             //Try reconnection after a wait time
             #statIterator := 0;
             #statState.connection := #STATE_WAIT;
           END_IF;
         END_IF;
         //Job completed without error
       ELSIF (#instTCON.DONE) THEN

         //Connection successfully established
         #diagnostics.statistics.totalReconnects := #diagnostics.statistics.totalReconnects + 1;
         #statState.connection := #OPERATION;

         #error := FALSE;

         //Reset all state machines
         #statState.receiver := #READ;
         #statState.sender := #STATE_INACTIVE;
         #statState.comReceiver := #LCOM_EXPECTED;
         #statState.comSender := #STATE_INACTIVE;
         //Receive
         #statReceive.trcvFct.dataOffset := 0;
         #statReceive.trcvFct.dataLength := 0;
         #statReceive.trcvFct.dataLengthRest := 0;
         #statReceive.trcvFct.dataReceived := FALSE;
         #statReceive.tempTelegram.index := 0;
         #statReceive.tempTelegram.telegramType := 0;
         #statReceive.numberOfLComHeader := 0;
         #statReceive.dataTelegram.totalMessageLength := 0;
         #statReceive.dataTelegram.actPackageLength := 0;
         #statReceive.dataTelegram.ackMessageOffset := 0;
         #statReceive.dataTelegram.messageOffset := 0;
         #statReceive.dataTelegram.ackMessageCounter := 0;
         #statReceive.dataTelegram.messageCounter := 0;
         #statReceive.userData.totalLength := 0;
         #statReceive.userData.offset := 0;
         //Send
         #statSend.tsendFct.dataLengthRest := 0;
         #statSend.tsendFct.dataOffset := 0;
         #statSend.tsendFct.status := 16#0000;
         #statSend.expectedAck.package1.offset := 0;
         #statSend.dataTelegram.messageCounter := 0;
         #statSend.dataTelegram.ackMessageCounter := 0;
         #statSend.dataTelegram.messageOffset := 0;
         #statSend.dataTelegram.ackMessageOffset := 0;
         #statSend.dataTelegram.actPackageLength := 0;
         #statSend.dataTelegram.totalMessageLength := 0;
         #statSend.numberOfLComPackage := 0;
         #statSend.userData.totalLength := 0;
         #statSend.userData.offset := 0;
         #statSend.userData.sendCycleViolation := FALSE;
         #statOldSend := FALSE;

         #diagnostics.statistics.maxMsgSendingTime := T#0ms;
         #diagnostics.localConfig.sender.cycleTime := T#0ms;
         #diagnostics.localConfig.sender.ackTimeout := T#0ms;

         #diagnostics.statistics.lastTimeSync.YEAR := 2200;
         #statCopyNBytes := 0;

         //Reset all timer
         #instLocalLifeSignCycleTimer(IN := FALSE,
                                      PT := #diagnostics.localConfig.connection.lifeSignCycleTime);

         #instPartnerLifeSignCycleTimer(IN := FALSE,
                                        PT := (#diagnostics.partnerConfig.connnection.lifeSignCycleTime));

         #instLocalCycleTimeTimer(IN := FALSE,
                                  PT := #diagnostics.localConfig.sender.cycleTime);

         #instExpectedAckPackage1(IN := FALSE,
                                  PT := #diagnostics.localConfig.sender.ackTimeout);

         #instSyncTimer(IN := FALSE,
                        PT := T#1s);

         #instSendErrorTimer(IN := FALSE,
                             PT := #MAX_TRIAL_TIME);

         #instRcvErrorTimer(IN := FALSE,
                            PT := #MAX_TRIAL_TIME);

         //Reset all active failures in the diagnostics buffer
         FOR #statIterator := 0 TO #DIAG_BUFFER_UPPER_LIM BY 1 DO
           #diagnostics.buffer[#statIterator].isActive := FALSE;
         END_FOR;

         //With LCom protocol
         IF (#diagnostics.localConfig.connection.useLComProtocol = TRUE) THEN

           IF (#statConnectAttempts MOD 2 = 0) THEN
             //1st try LCom Version 2.0
             #statActualLocalLComVersion := #LCOM_HEADER_V2;
             #statSend.configTelegramV2.LComVersion := #LCOM_HEADER_V2;
             #statSend.configTelegramV2.status := BOOL_TO_BYTE(#diagnostics.localConfig.timeSync.usePartnerTimestamps);
             #statSend.configTelegramV2.sendModeSyncTime := #diagnostics.localConfig.timeSync.sendMode;
             #statSend.configTelegramV2.lifeSignCycle := #diagnostics.localConfig.connection.lifeSignCycleTime;
             #statSend.configTelegramV2.cycleTime := #configuration.sender.cycleTime;
             #statSend.configTelegramV2.ackTimeOut := #configuration.sender.ackTimeout;
             #statSend.configTelegramV2.maxSendDataLength := #diagnostics.localConfig.sizeOfSendBuffer;
             #statSend.configTelegramV2.maxReceiveDataLength := #diagnostics.localConfig.sizeOfReceiveBuffer;

             #statSend.dataTelegram.LComVersion := #statSend.configTelegramV2.LComVersion;
           ELSE
             //2nd try LCom Version 1.0
             #statActualLocalLComVersion := #LCOM_HEADER_V1;
             #statSend.configTelegramV1.LComVersion := #LCOM_HEADER_V1;
             #statSend.configTelegramV1.comMode := 16#03;
             #statSend.configTelegramV1.slidingWindow := 1;
             #statSend.configTelegramV1.status := BOOL_TO_BYTE(#diagnostics.localConfig.timeSync.usePartnerTimestamps);
             #statSend.configTelegramV1.sendModeSyncTime := #diagnostics.localConfig.timeSync.sendMode;

             #statSend.dataTelegram.LComVersion := #statSend.configTelegramV1.LComVersion;

             //Check max. lifeSignCycleTime
             IF (#diagnostics.localConfig.connection.lifeSignCycleTime > T#65535ms) THEN

               #statDiag.bufferIndex := #statDiag.bufferIndex + 1;
               #statDiag.buffer[#statDiag.bufferIndex].additionalValue4 := #diagnostics.localConfig.connection.lifeSignCycleTime;
               #diagnostics.localConfig.connection.lifeSignCycleTime := T#65535ms;

               #statDiag.buffer[#statDiag.bufferIndex].status := "LCOM_WARN_LIFE_SIGN_LIMITATION";
               #statDiag.buffer[#statDiag.bufferIndex].subFunctionErrorID := 16#0000;
               #statDiag.buffer[#statDiag.bufferIndex].additionalValue1 := 65535.0;
               #statDiag.buffer[#statDiag.bufferIndex].additionalValue2 := 0.0;
               #statDiag.buffer[#statDiag.bufferIndex].additionalValue3 := 0.0;
             ELSE
               ;
             END_IF;
             #statSend.configTelegramV1.lifeSignCycle := TIME_TO_UINT(#diagnostics.localConfig.connection.lifeSignCycleTime);

             //Check max.sizeOfSendBuffer
             IF (#diagnostics.localConfig.sizeOfSendBuffer > 65535) THEN
               #diagnostics.localConfig.sizeOfSendBuffer := 65535;
               #statSend.configTelegramV1.maxSendDataLength := 65535;
             ELSE
               #statSend.configTelegramV1.maxSendDataLength := UDINT_TO_UINT(#diagnostics.localConfig.sizeOfSendBuffer);
             END_IF;

             //Check max.sizeOfReceiveBuffer
             IF (#diagnostics.localConfig.sizeOfReceiveBuffer > 65535) THEN
               #diagnostics.localConfig.sizeOfReceiveBuffer := 65535;
               #statSend.configTelegramV1.maxReceiveDataLength := 65535;
             ELSE
               #statSend.configTelegramV1.maxReceiveDataLength := UDINT_TO_UINT(#diagnostics.localConfig.sizeOfReceiveBuffer);
             END_IF;

           END_IF;
           //Set telegram type of data telegrams for LCom Version 1.0 and 2.0
           #statSend.dataTelegram.telegramType := 16#0A;

           //Start sender config directly with LCom protocol
           #statState.cfgSender := #STATE_INIT;
         ELSE
           //without LCom
           #statCompare.sender.cycleTime := #configuration.sender.cycleTime;
           #diagnostics.localConfig.sender.cycleTime := #configuration.sender.cycleTime;

           #diagnostics.partnerConfig.sizeOfReceiveBuffer := 0;
           #diagnostics.partnerConfig.sizeOfSendBuffer := 0;
           #connected := TRUE;
           #statState.cfgSender := #OPERATION;

           #statDiag.bufferIndex := #statDiag.bufferIndex + 1;
           #statDiag.buffer[#statDiag.bufferIndex].status := "LCOM_STATUS_TCP_CONNECTED";
           #statDiag.buffer[#statDiag.bufferIndex].subFunctionErrorID := 16#0000;
           #statDiag.buffer[#statDiag.bufferIndex].additionalValue1 := 0.0;
           #statDiag.buffer[#statDiag.bufferIndex].additionalValue2 := 0.0;
           #statDiag.buffer[#statDiag.bufferIndex].additionalValue3 := 0.0;
           #statDiag.buffer[#statDiag.bufferIndex].additionalValue4 := T#0ms;
         END_IF;
         //TCON still in progress
       ELSE
         IF (#diagnostics.localConfig.connection.isClient) THEN

           #statDiag.bufferIndex := #statDiag.bufferIndex + 1;
           #statDiag.buffer[#statDiag.bufferIndex].status := "LCOM_STATUS_CLIENT_TRY_CONNECT";
           #statDiag.buffer[#statDiag.bufferIndex].subFunctionErrorID := 16#0000;
           #statDiag.buffer[#statDiag.bufferIndex].additionalValue1 := 0.0;
           #statDiag.buffer[#statDiag.bufferIndex].additionalValue2 := 0.0;
           #statDiag.buffer[#statDiag.bufferIndex].additionalValue3 := 0.0;
           #statDiag.buffer[#statDiag.bufferIndex].additionalValue4 := T#0ms;
         ELSE
           #statDiag.bufferIndex := #statDiag.bufferIndex + 1;
           #statDiag.buffer[#statDiag.bufferIndex].status := "LCOM_STATUS_SERVER_PORT_OPEN";
           #statDiag.buffer[#statDiag.bufferIndex].subFunctionErrorID := 16#0000;
           #statDiag.buffer[#statDiag.bufferIndex].additionalValue1 := 0.0;
           #statDiag.buffer[#statDiag.bufferIndex].additionalValue2 := 0.0;
           #statDiag.buffer[#statDiag.bufferIndex].additionalValue3 := 0.0;
           #statDiag.buffer[#statDiag.bufferIndex].additionalValue4 := T#0ms;
         END_IF;
       END_IF;

     #STATE_WAIT:

       //Wait and then establish the connection
       IF (#statIterator > #STATE_WAIT) THEN

         #instTCON(REQ := FALSE,
                   ID := #configuration.connection.connectionID,
                   CONNECT := #statTconPar);

         #instTSEND(REQ := FALSE,
                    ID := #statTconPar.ID,
                    DATA := #statSend.tsendFct.data);

         #instTRCV(EN_R := FALSE,
                   ID := #statTconPar.ID,
                   DATA := #statReceive.trcvFct.data);

         #instTDISCON(REQ := FALSE,
                      ID := #statTconPar.ID);

         IF (#diagnostics.localConfig.connection.isClient) THEN
           #statState.connection := #OPEN_CLIENT;
           #statTconPar.ActiveEstablished := TRUE;
         ELSE
           #statState.connection := #OPEN_SERVER;
           #statTconPar.ActiveEstablished := FALSE;
         END_IF;

       ELSE
         #statIterator := #statIterator + 1;
       END_IF;

     #FINISH_TSEND:

       IF (#statIterator > #STATE_WAIT) THEN
         #statIterator := 0;
         #statState.connection := #FINISH_TRCV;
       ELSE
         #instTSEND(REQ := TRUE,
                    LEN := #statSend.tsendFct.dataOffset,
                    ID := #statTconPar.ID,
                    DATA := #statSend.tsendFct.data,
                    STATUS => #statSend.tsendFct.status);

         IF ((#statSend.tsendFct.status = 16#0000) OR (#instTSEND.ERROR)) THEN
           //"TSEND" instruction is finished
           #statState.connection := #FINISH_TRCV;
         ELSE
           ;//"TSEND" instruction still in process
         END_IF;
       END_IF;
       #statIterator := #statIterator + 1;
     #FINISH_TRCV:

       IF (#statIterator > #STATE_WAIT) THEN
         #statState.connection := #CALL_TDISCON;
       ELSE
         #instTRCV(EN_R := TRUE,
                   ID := #diagnostics.localConfig.connection.connectionID,
                   LEN := 0,
                   ADHOC := TRUE,
                   NDR => #statReceive.trcvFct.dataReceived,
                   RCVD_LEN => #statReceive.trcvFct.dataLength,
                   DATA := #statReceive.trcvFct.data);

         //Is the "TRCV" instruction still in process
         IF (#instTRCV.ERROR OR NOT #instTRCV.BUSY) THEN
           #statState.connection := #CALL_TDISCON;
         ELSE
           ;//TRCV instruction still in process
         END_IF;
       END_IF;
       #statIterator := #statIterator + 1;

     #CLOSE_CONNECTION:

       //reset FB Outputs
       #connected := FALSE;
       #sending := FALSE;
       #receivedDataLength := 0;
       #error := FALSE;

       //Is "TSEND" instruction still in process ?
       IF (#statSend.tsendFct.status <> 16#0000) THEN
         //"TSEND" instruction still in process
         #statState.connection := #FINISH_TSEND;
         #statIterator := 0;
       ELSE
         ;//"TSEND" instruction is finished
       END_IF;

       #instTRCV(EN_R := TRUE,
                 ID := #diagnostics.localConfig.connection.connectionID,
                 LEN := 0,
                 ADHOC := TRUE,
                 NDR => #statReceive.trcvFct.dataReceived,
                 RCVD_LEN => #statReceive.trcvFct.dataLength,
                 DATA := #statReceive.trcvFct.data);

       //Is the "TRCV" instruction still in process
       IF (#instTRCV.ERROR OR NOT #instTRCV.BUSY) THEN
         #statState.connection := #CALL_TDISCON;
       ELSE
         #statState.connection := #FINISH_TRCV;
         #statIterator := 0;
       END_IF;

     #CALL_TDISCON:

       #instTSEND(REQ := FALSE,
                  LEN := #statSend.tsendFct.dataOffset,
                  ID := #statTconPar.ID,
                  DATA := #statSend.tsendFct.data);

       #instTRCV(EN_R := FALSE,
                 ID := #diagnostics.localConfig.connection.connectionID,
                 LEN := 0,
                 ADHOC := TRUE,
                 NDR => #statReceive.trcvFct.dataReceived,
                 RCVD_LEN => #statReceive.trcvFct.dataLength,
                 DATA := #statReceive.trcvFct.data);

       #instTDISCON(REQ := TRUE,
                    ID := #statTconPar.ID);

       //Error occurred during processing
       IF (#instTDISCON.ERROR) THEN

         #statDiag.bufferIndex := #statDiag.bufferIndex + 1;
         #statDiag.buffer[#statDiag.bufferIndex].status := "LCOM_ERR_CLOSE_CONNECTION";
         #statDiag.buffer[#statDiag.bufferIndex].subFunctionErrorID := #instTDISCON.STATUS;
         #statDiag.buffer[#statDiag.bufferIndex].additionalValue1 := 0.0;
         #statDiag.buffer[#statDiag.bufferIndex].additionalValue2 := 0.0;
         #statDiag.buffer[#statDiag.bufferIndex].additionalValue3 := 0.0;
         #statDiag.buffer[#statDiag.bufferIndex].additionalValue4 := T#0ms;

         #statState.connection := #STATE_INACTIVE_PREPARE;

         #instTDISCON(REQ := FALSE,
                      ID := #statTconPar.ID);

       ELSIF (#instTDISCON.DONE) THEN

         #instTDISCON(REQ := FALSE,
                      ID := #statTconPar.ID);
         //Job executed without errors
         IF (#enable AND (NOT #statFallingEdgeEnable)) THEN
           //Reconnect automatically if not in disconnecting process
           #statIterator := 0;
           #statState.connection := #STATE_WAIT;
         ELSE
           //Reset all active failures in the diagnostics buffer
           FOR #statIterator := 0 TO #DIAG_BUFFER_UPPER_LIM BY 1 DO
             #diagnostics.buffer[#statIterator].isActive := FALSE;
           END_FOR;

           #statState.connection := #STATE_INACTIVE_PREPARE;
         END_IF;
         //Job is not completed yet
       ELSE
         ;//Wait until job is finished
       END_IF;
     #ERROR_STATE:
       ;

   END_CASE;

   // -----------------------------------------------------------------------------------------------------------
   //Diagnostics buffer
   // -----------------------------------------------------------------------------------------------------------
   diag:
   //Diagnostics entry is in the temp. buffer
   IF (#statDiag.bufferIndex <> 255) THEN

     //Get current time
     #statRet := RD_LOC_T(#tempActTime);
     //init
     #statDiag.actualIndex := 0;

     WHILE (#statDiag.actualIndex <= #statDiag.bufferIndex) DO

       #tempUDint := 0;
       //Check if the failure is already in the buffer and still active
       FOR #statIterator := 0 TO #DIAG_BUFFER_UPPER_LIM BY 1 DO

         IF (#diagnostics.buffer[#statIterator].isActive = TRUE) THEN

           IF ((#statDiag.buffer[#statDiag.actualIndex].status = "LCOM_WARN_SEND_CYCLE_EXPIRED")
             AND
             (#diagnostics.buffer[#statIterator].status = "LCOM_WARN_SEND_CYCLE_EXPIRED")
             AND
             (#diagnostics.buffer[#statIterator].additionalValue1 = #statDiag.buffer[#statDiag.actualIndex].additionalValue1)
             AND
             (#diagnostics.buffer[#statIterator].additionalValue2 = #statDiag.buffer[#statDiag.actualIndex].additionalValue2)
             AND
             (#diagnostics.buffer[#statIterator].additionalValue3 = #statDiag.buffer[#statDiag.actualIndex].additionalValue3)) THEN
             //Retrigger just the activation time
             #diagnostics.buffer[#statIterator].timestamp := #tempActTime;
             #diagnostics.buffer[#statIterator].additionalValue4 := #statDiag.buffer[#statDiag.actualIndex].additionalValue4;
             #tempUDint := 100;
             EXIT;
           ELSIF ((#diagnostics.buffer[#statIterator].status = #statDiag.buffer[#statDiag.actualIndex].status)
             AND
             (#diagnostics.buffer[#statIterator].additionalValue1 = #statDiag.buffer[#statDiag.actualIndex].additionalValue1)
             AND
             (#diagnostics.buffer[#statIterator].additionalValue2 = #statDiag.buffer[#statDiag.actualIndex].additionalValue2)
             AND
             (#diagnostics.buffer[#statIterator].additionalValue3 = #statDiag.buffer[#statDiag.actualIndex].additionalValue3)
             AND
             (#diagnostics.buffer[#statIterator].additionalValue4 = #statDiag.buffer[#statDiag.actualIndex].additionalValue4)) THEN
             //Retrigger just the activation time
             #diagnostics.buffer[#statIterator].timestamp := #tempActTime;
             #tempUDint := 100;
             EXIT;
           ELSE
             ;//ErrorId is not in the diagnostics buffer
           END_IF;
         END_IF;
       END_FOR;

       IF (#tempUDint = 100) THEN
         ;//ErrorId was already retriggered
       ELSE
         //Check range of diagnostics ring buffer [0...LCOM_DIAG_ARRAY]
           IF ((#diagnostics.bufferIndex = 255) OR (#diagnostics.bufferIndex = #DIAG_BUFFER_UPPER_LIM)) THEN
           #diagnostics.bufferIndex := 0;
         ELSE
           #diagnostics.bufferIndex := #diagnostics.bufferIndex + 1;
         END_IF;

         //Stored new entry in the diagnostics buffer
         #diagnostics.buffer[#diagnostics.bufferIndex].status := #statDiag.buffer[#statDiag.actualIndex].status;
         #diagnostics.buffer[#diagnostics.bufferIndex].timestamp := #tempActTime;
         #diagnostics.buffer[#diagnostics.bufferIndex].isActive := TRUE;

         #diagnostics.buffer[#diagnostics.bufferIndex].subFunctionErrorID := #statDiag.buffer[#statDiag.actualIndex].subFunctionErrorID;
         #diagnostics.buffer[#diagnostics.bufferIndex].additionalValue1 := #statDiag.buffer[#statDiag.actualIndex].additionalValue1;
         #diagnostics.buffer[#diagnostics.bufferIndex].additionalValue2 := #statDiag.buffer[#statDiag.actualIndex].additionalValue2;
         #diagnostics.buffer[#diagnostics.bufferIndex].additionalValue3 := #statDiag.buffer[#statDiag.actualIndex].additionalValue3;
         #diagnostics.buffer[#diagnostics.bufferIndex].additionalValue4 := #statDiag.buffer[#statDiag.actualIndex].additionalValue4;
       END_IF;

       IF ((#diagnostics.buffer[#diagnostics.bufferIndex].status = "LCOM_STATUS_TCP_CONNECTED")
         OR (#diagnostics.buffer[#diagnostics.bufferIndex].status = "LCOM_STATUS_LCOM_CONNECTED_V1")
         OR (#diagnostics.buffer[#diagnostics.bufferIndex].status = "LCOM_STATUS_LCOM_CONNECTED_V2"))
       THEN
         #statConnectAttempts := 0;
         #diagnostics.statistics.lastConnect := #tempActTime;
       END_IF;

       //Set FB status
       #status := #statDiag.buffer[#statDiag.actualIndex].status;

       //Check if FB.error has been set ?
       IF ((#statDiag.buffer[#statDiag.actualIndex].status >= "LCOM_ERR_COM_SERVICE")//16#8200
         AND
         (#statDiag.buffer[#statDiag.actualIndex].status <= "LCOM_ERR_WRONG_TELEGRAM_ID"))//16#8614
       THEN

         #error := TRUE;
         #connected := FALSE;
         #sending := FALSE;
         #dataReceived := FALSE;
         #receivedDataLength := 0;

         //Check if FB.busy has been set ?
         IF ((#statDiag.buffer[#statDiag.actualIndex].status >= "LCOM_ERR_OPEN_CLIENT")//16#8600
           AND
           (#statDiag.buffer[#statDiag.actualIndex].status <= "LCOM_ERR_WRONG_TELEGRAM_ID"))//16#8614
         THEN
           #busy := TRUE;
         ELSE
           #busy := FALSE;
         END_IF;

         EXIT;//Leave loop
       ELSE
         ;
       END_IF;

       //Increase index
       #statDiag.actualIndex := #statDiag.actualIndex + 1;

     END_WHILE;
   ELSE
     ;//No failure
   END_IF;//End: Diagnostics buffer
END_FUNCTION_BLOCK

FUNCTION "ResetFaults" : Void   // FC1, FBD
{ S7_Optimized_Access := 'TRUE' }
VERSION : 0.1
   VAR_OUTPUT
      NoReadFault : Bool;
      "Mis-MatchFault" : Bool;
      "Mis-TriggerFault" : Bool;
   END_VAR
BEGIN

REGION Network 1 (SCL)

       #NoReadFault := 0;
       #"Mis-MatchFault" := 0;
       #"Mis-TriggerFault" := 0;
END_REGION
END_FUNCTION

FUNCTION "ToSPC" : Void   // FC2, FBD
{ S7_Optimized_Access := 'TRUE' }
VERSION : 0.1
   VAR_INPUT
      NoReadFault : Bool;
      MisMatchFault : Bool;
      MisTriggerFauld : Bool;
      ValidMaterialNumber : Bool;
      EnigmaDisable : Bool;
   END_VAR
   VAR_OUTPUT
      NoReadFaultToSPC : Bool;
      MisMatchFaultToSPC : Bool;
      MisTriggerFauldToSPC : Bool;
      ValidMaterialNumberToSPC : Bool;
      EnigmaDisableToSPC : Bool;
   END_VAR
BEGIN

REGION Network 1
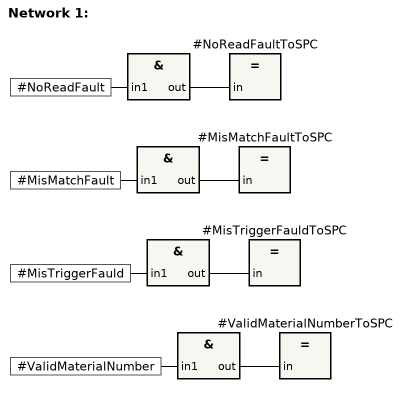
   #NoReadFaultToSPC := #NoReadFault;
   #MisMatchFaultToSPC := #MisMatchFault;
   #MisTriggerFauldToSPC := #MisTriggerFauld;
   #ValidMaterialNumberToSPC := #ValidMaterialNumber;
END_REGION
END_FUNCTION

FUNCTION "LightsStatus" : Void   // FC3, LAD
{ S7_Optimized_Access := 'TRUE' }
VERSION : 0.1
BEGIN

REGION Network 1: Lable istic vypnuty
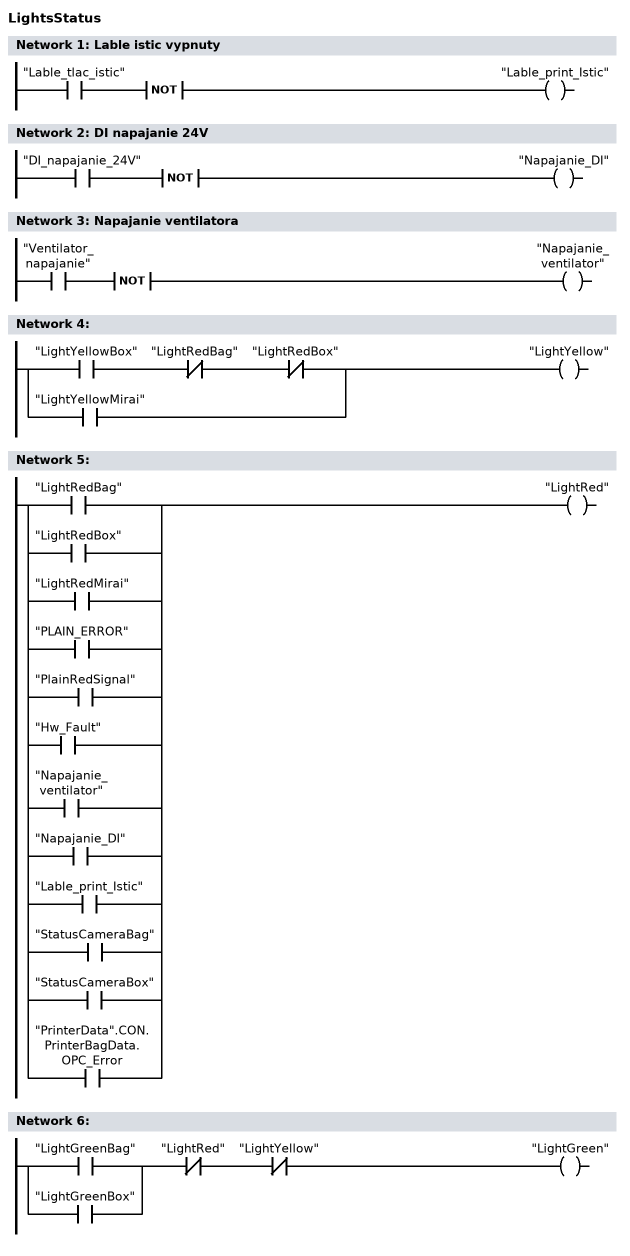
   RUNG wire#powerrail
      Contact( "Lable_tlac_istic" )
      Not()
      Coil( "Lable_print_Istic" )
   END_RUNG
   // the same network as SCL:
   "Lable_print_Istic" := NOT "Lable_tlac_istic";
END_REGION

REGION Network 2: DI napajanie 24V
   RUNG wire#powerrail
      Contact( "DI_napajanie_24V" )
      Not()
      Coil( "Napajanie_DI" )
   END_RUNG
   // the same network as SCL:
   "Napajanie_DI" := NOT "DI_napajanie_24V";
END_REGION

REGION Network 3: Napajanie ventilatora
   RUNG wire#powerrail
      Contact( "Ventilator_napajanie" )
      Not()
      Coil( "Napajanie_ventilator" )
   END_RUNG
   // the same network as SCL:
   "Napajanie_ventilator" := NOT "Ventilator_napajanie";
END_REGION

REGION Network 4
   RUNG wire#powerrail
      Contact( "LightYellowBox" )
      I_Contact( "LightRedBag" )
      I_Contact( "LightRedBox" )
      wire#w1
      Coil( "LightYellow" )
   END_RUNG
   RUNG wire#powerrail
      Contact( "LightYellowMirai" )
   END_RUNG wire#w1
   // the same network as SCL:
   "LightYellow" := ("LightYellowBox" AND NOT "LightRedBag" AND NOT "LightRedBox") OR "LightYellowMirai";
END_REGION

REGION Network 5
   RUNG wire#powerrail
      Contact( "LightRedBag" )
      wire#w1
      Coil( "LightRed" )
   END_RUNG
   RUNG wire#powerrail
      Contact( "LightRedBox" )
   END_RUNG wire#w1
   RUNG wire#powerrail
      Contact( "LightRedMirai" )
   END_RUNG wire#w1
   RUNG wire#powerrail
      Contact( "PLAIN_ERROR" )
   END_RUNG wire#w1
   RUNG wire#powerrail
      Contact( "PlainRedSignal" )
   END_RUNG wire#w1
   RUNG wire#powerrail
      Contact( "Hw_Fault" )
   END_RUNG wire#w1
   RUNG wire#powerrail
      Contact( "Napajanie_ventilator" )
   END_RUNG wire#w1
   RUNG wire#powerrail
      Contact( "Napajanie_DI" )
   END_RUNG wire#w1
   RUNG wire#powerrail
      Contact( "Lable_print_Istic" )
   END_RUNG wire#w1
   RUNG wire#powerrail
      Contact( "StatusCameraBag" )
   END_RUNG wire#w1
   RUNG wire#powerrail
      Contact( "StatusCameraBox" )
   END_RUNG wire#w1
   RUNG wire#powerrail
      Contact( "PrinterData".CON.PrinterBagData.OPC_Error )
   END_RUNG wire#w1
   // the same network as SCL:
   "LightRed" := "LightRedBag" OR "LightRedBox" OR "LightRedMirai" OR "PLAIN_ERROR" OR "PlainRedSignal" OR "Hw_Fault" OR "Napajanie_ventilator" OR "Napajanie_DI" OR "Lable_print_Istic" OR "StatusCameraBag" OR "StatusCameraBox" OR "PrinterData".CON.PrinterBagData.OPC_Error;
END_REGION

REGION Network 6
   RUNG wire#powerrail
      Contact( "LightGreenBag" )
      wire#w1
      I_Contact( "LightRed" )
      I_Contact( "LightYellow" )
      Coil( "LightGreen" )
   END_RUNG
   RUNG wire#powerrail
      Contact( "LightGreenBox" )
   END_RUNG wire#w1
   // the same network as SCL:
   "LightGreen" := ("LightGreenBag" OR "LightGreenBox") AND NOT "LightRed" AND NOT "LightYellow";
END_REGION
END_FUNCTION

FUNCTION "TimeServerCom" : Void   // FC4, LAD
{ S7_Optimized_Access := 'TRUE' }
VERSION : 0.1
   VAR_INPUT
      BatchEndTime : String;
   END_VAR
   VAR_OUTPUT
      "Date" : String;
      "Time" : String;
      BatchStatus : Byte;
   END_VAR
   VAR_TEMP
      ReturnVal : Int;
      DateTime : DTL;
      y : String;
      mo : String;
      d : String;
      h : String;
      "m" : String;
      s : String;
      Dummy1 : UInt;
      BatchDayEnd : Int;
      BatchMinuteEnd : Int;
      i : Int;
      year : Array[0..3] of Char;
      month : Array[0..1] of Char;
      day : Array[0..1] of Char;
      hour : Array[0..1] of Char;
      minute : Array[0..1] of Char;
      second : Array[0..1] of Char;
      Date1 : String;
      Time1 : String;
      index1 : Int;
      DayOPC : Int;
      MonthOPC : Int;
      YearOPC : Int;
      HourOPC : Int;
      MinuteOPC : Int;
      BatchDummy1 : String;
   END_VAR
   VAR CONSTANT
      WarningBatch : Time := T#2H;
      ErrorBatch : Time := T#10M;
   END_VAR
BEGIN

REGION Network 1 (SCL)
   REGION TimeDate
       // Read time and date and convert it to string
       #ReturnVal := RD_LOC_T(#DateTime);
       //convert time and data to the seprate string
       VAL_STRG(IN := #DateTime.YEAR,
                SIZE := 4,
                PREC := 0,
                FORMAT := 0,
                P := 1,
                OUT => #y);
       //month
       VAL_STRG(IN := #DateTime.MONTH,
                SIZE := 2,
                PREC := 0,
                FORMAT := 0,
                P := 1,
                OUT => #mo);
       //day
       VAL_STRG(IN := #DateTime.DAY,
                SIZE := 2,
                PREC := 0,
                FORMAT := 0,
                P := 1,
                OUT => #d);
       //hour
       VAL_STRG(IN := #DateTime.HOUR,
                SIZE := 2,
                PREC := 0,
                FORMAT := 0,
                P := 1,
                OUT => #h);
       //minute
       VAL_STRG(IN := #DateTime.MINUTE,
                SIZE := 2,
                PREC := 0,
                FORMAT := 0,
                P := 1,
                OUT => #m);
       //second
       VAL_STRG(IN := #DateTime.SECOND,
                SIZE := 2,
                PREC := 0,
                FORMAT := 0,
                P := 1,
                OUT => #s);
   END_REGION
   REGION toChar
       // change the string to char
       //year
       Strg_TO_Chars(Strg := #y,
                     pChars := 0,
                     Cnt => #Dummy1,
                     Chars := #year);
       //month
       Strg_TO_Chars(Strg := #mo,
                     pChars := 0,
                     Cnt => #Dummy1,
                     Chars := #month);
       //day
       Strg_TO_Chars(Strg := #d,
                     pChars := 0,
                     Cnt => #Dummy1,
                     Chars := #day);
       //hour
       Strg_TO_Chars(Strg := #h,
                     pChars := 0,
                     Cnt => #Dummy1,
                     Chars := #hour);
         //minute
       Strg_TO_Chars(Strg := #m,
                     pChars := 0,
                     Cnt => #Dummy1,
                     Chars := #minute);
       Strg_TO_Chars(Strg := #s,
                     pChars := 0,
                     Cnt => #Dummy1,
                     Chars := #second);
   END_REGION
   REGION NullChar
       // check for null char and replace it with zero
       //year
       FOR #i := 0 TO 3 DO
           IF #year[#i] = ' '
           THEN
               #year[#i] := '0';
           END_IF;
       END_FOR;
       //month
       FOR #i := 0 TO 1 DO
           IF #month[#i] = ' '
           THEN
               #month[#i] := '0';
           END_IF;
       END_FOR;
       //day
       FOR #i := 0 TO 1 DO
           IF #day[#i] = ' '
           THEN
               #day[#i] := '0';
           END_IF;
       END_FOR;
       //hour
       FOR #i := 0 TO 1 DO
           IF #hour[#i] = ' '
           THEN
               #hour[#i] := '0';
           END_IF;
       END_FOR;
       //minute
       FOR #i := 0 TO 1 DO
           IF #minute[#i] = ' '
           THEN
               #minute[#i] := '0';
           END_IF;
       END_FOR;
       //second
       FOR #i := 0 TO 1 DO
           IF #second[#i] = ' '
           THEN
               #second[#i] := '0';
           END_IF;
       END_FOR;
   END_REGION
   REGION Output
       // Time and date as a string
       Chars_TO_Strg(Chars := #year,
                     pChars := 0,
                     Cnt := 4,
                     Strg => #y);
       Chars_TO_Strg(Chars := #month,
                     pChars := 0,
                     Cnt := 2,
                     Strg => #mo);
       Chars_TO_Strg(Chars := #day,
                     pChars := 0,
                     Cnt := 2,
                     Strg => #d);
       Chars_TO_Strg(Chars := #hour,
                     pChars := 0,
                     Cnt := 2,
                     Strg => #h);
       Chars_TO_Strg(Chars := #minute,
                     pChars := 0,
                     Cnt := 2,
                     Strg => #m);
       Chars_TO_Strg(Chars := #second,
                     pChars := 0,
                     Cnt := 2,
                     Strg => #s);
       #Date1 := CONCAT(IN1 := #y, IN2 := #mo);
       #Date := CONCAT(IN1 := #Date1, IN2 := #d);
       #Time1 := CONCAT(IN1 := #h, IN2 := #m);
       #Time := CONCAT(IN1 := #Time1, IN2 := #s);
   END_REGION
   REGION Batch
       // Creat the alarm and error for the planed batch end time
       // day
       #index1 := FIND(IN1 := #BatchEndTime, IN2 := '/');
       STRG_VAL(IN:=#BatchEndTime,
                FORMAT:=0,
                P:=1,
                OUT=>#DayOPC);
       #BatchDummy1:= DELETE(IN:=#BatchEndTime, L:=#index1, P:=1);
       //month
       #index1 := FIND(IN1 := #BatchDummy1, IN2 := '/');
       STRG_VAL(IN := #BatchDummy1,
                FORMAT := 0,
                P := 1,
                OUT => #MonthOPC);
       #BatchDummy1 := DELETE(IN := #BatchDummy1, L := #index1, P := 1);
       //year
       #index1 := FIND(IN1 := #BatchDummy1, IN2 := ' ');
       STRG_VAL(IN := #BatchDummy1,
                FORMAT := 0,
                P := 1,
                OUT => #YearOPC);
       #BatchDummy1 := DELETE(IN := #BatchDummy1, L := #index1, P := 1);
       //hour
       #index1 := FIND(IN1 := #BatchDummy1, IN2 := ':');
       STRG_VAL(IN := #BatchDummy1,
                FORMAT := 0,
                P := 1,
                OUT => #HourOPC);
       #BatchDummy1 := DELETE(IN := #BatchDummy1, L := #index1, P := 1);
       //minute
       #index1 := FIND(IN1 := #BatchDummy1, IN2 := ':');
       STRG_VAL(IN := #BatchDummy1,
                FORMAT := 0,
                P := 1,
                OUT => #MinuteOPC);
       #BatchDayEnd:= (#YearOPC - #DateTime.YEAR)*365+(#MonthOPC - #DateTime.MONTH)*30+( #DayOPC - #DateTime.DAY);
       #BatchMinuteEnd := (#HourOPC - #DateTime.HOUR) * 60 + (#MinuteOPC - #DateTime.MINUTE);

       IF #BatchDayEnd = 0 THEN
           IF #BatchMinuteEnd < 60 AND #BatchMinuteEnd > 11 THEN
               #BatchStatus := 1; //warning
           ELSIF #BatchMinuteEnd <= 11 AND #BatchMinuteEnd >0 THEN
               #BatchStatus := 2;//batch error
           ELSIF #BatchMinuteEnd = 0 THEN 
               #BatchStatus := 3;
           ELSIF #BatchMinuteEnd <0 THEN
               #BatchStatus := 3;
               ELSE
               #BatchStatus := 0;
           END_IF;
       ELSIF  #BatchDayEnd < 0  THEN
           #BatchStatus := 3;
       ELSE
           #BatchStatus := 0;
       END_IF;
   END_REGION
END_REGION
END_FUNCTION

FUNCTION "Counter_32Bit_1" : Void   // FC5, FBD
{ S7_Optimized_Access := 'TRUE' }
VERSION : 0.1
   VAR_INPUT
      Varia : UDInt;
   END_VAR
   VAR_IN_OUT
      CountedValue : UDInt;
   END_VAR
   VAR_TEMP
      CountedValueDummy : UDInt;
   END_VAR
BEGIN

REGION Network 1 (SCL)
   #CountedValueDummy := #CountedValue;
   #CountedValueDummy := #CountedValueDummy + #Varia;
   #CountedValue := #CountedValueDummy;
END_REGION
END_FUNCTION

FUNCTION "HmiHandle" : Void   // FC6, LAD
{ S7_Optimized_Access := 'TRUE' }
VERSION : 0.1
   VAR_TEMP
      TmpS : String;
      TmpD : DInt;
   END_VAR
BEGIN

REGION Network 2